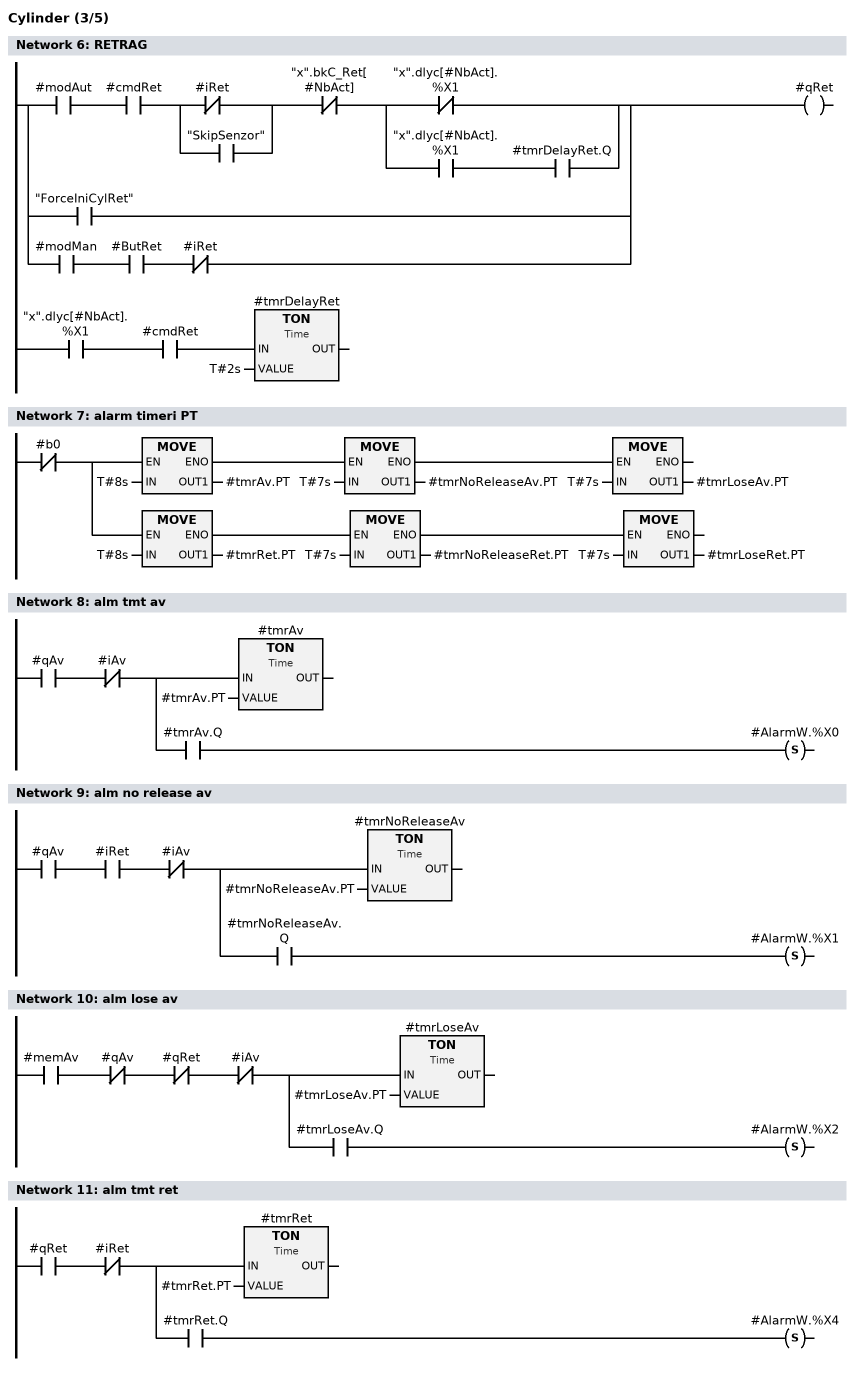
   #qRet := (#modAut AND #cmdRet AND (NOT #iRet OR "SkipSenzor") AND NOT "x".bkC_Ret[#NbAct] AND (NOT "x".dlyc[#NbAct].%X1 OR ("x".dlyc[#NbAct].%X1 AND #tmrDelayRet.Q))) OR "ForceIniCylRet" OR (#modMan AND #ButRet AND NOT #iRet);
   #tmrDelayRet.TON(IN := "x".dlyc[#NbAct].%X1 AND #cmdRet, PT := T#2s);   // TON coil
END_REGION

REGION Network 7: alarm timeri PT
   RUNG wire#powerrail
      I_Contact( #b0 )
      wire#w1
      Move(in := T#8s, out1 => #tmrAv.PT)
      Move(in := T#7s, out1 => #tmrNoReleaseAv.PT)
      Move(in := T#7s, out1 => #tmrLoseAv.PT)
   END_RUNG
   RUNG wire#w1
      Move(in := T#8s, out1 => #tmrRet.PT)
      Move(in := T#7s, out1 => #tmrNoReleaseRet.PT)
      Move(in := T#7s, out1 => #tmrLoseRet.PT)
   END_RUNG
   // the same network as SCL:
   IF NOT #b0 THEN
       #tmrAv.PT := T#8s;
       #tmrNoReleaseAv.PT := T#7s;
       #tmrLoseAv.PT := T#7s;
       #tmrRet.PT := T#8s;
       #tmrNoReleaseRet.PT := T#7s;
       #tmrLoseRet.PT := T#7s;
   END_IF;
END_REGION

REGION Network 8: alm tmt av
   #_w1 := #qAv AND NOT #iAv;
   #tmrAv.TON(IN := #_w1, PT := #tmrAv.PT);   // TON coil
   IF #_w1 AND #tmrAv.Q THEN #AlarmW.%X0 := TRUE; END_IF;
END_REGION

REGION Network 9: alm no release av
   #_w1 := #qAv AND #iRet AND NOT #iAv;
   #tmrNoReleaseAv.TON(IN := #_w1, PT := #tmrNoReleaseAv.PT);   // TON coil
   IF #_w1 AND #tmrNoReleaseAv.Q THEN #AlarmW.%X1 := TRUE; END_IF;
END_REGION

REGION Network 10: alm lose av
   #_w1 := #memAv AND NOT #qAv AND NOT #qRet AND NOT #iAv;
   #tmrLoseAv.TON(IN := #_w1, PT := #tmrLoseAv.PT);   // TON coil
   IF #_w1 AND #tmrLoseAv.Q THEN #AlarmW.%X2 := TRUE; END_IF;
END_REGION

REGION Network 11: alm tmt ret
   #_w1 := #qRet AND NOT #iRet;
   #tmrRet.TON(IN := #_w1, PT := #tmrRet.PT);   // TON coil
   IF #_w1 AND #tmrRet.Q THEN #AlarmW.%X4 := TRUE; END_IF;
END_REGION

REGION Network 12: alm no release ret
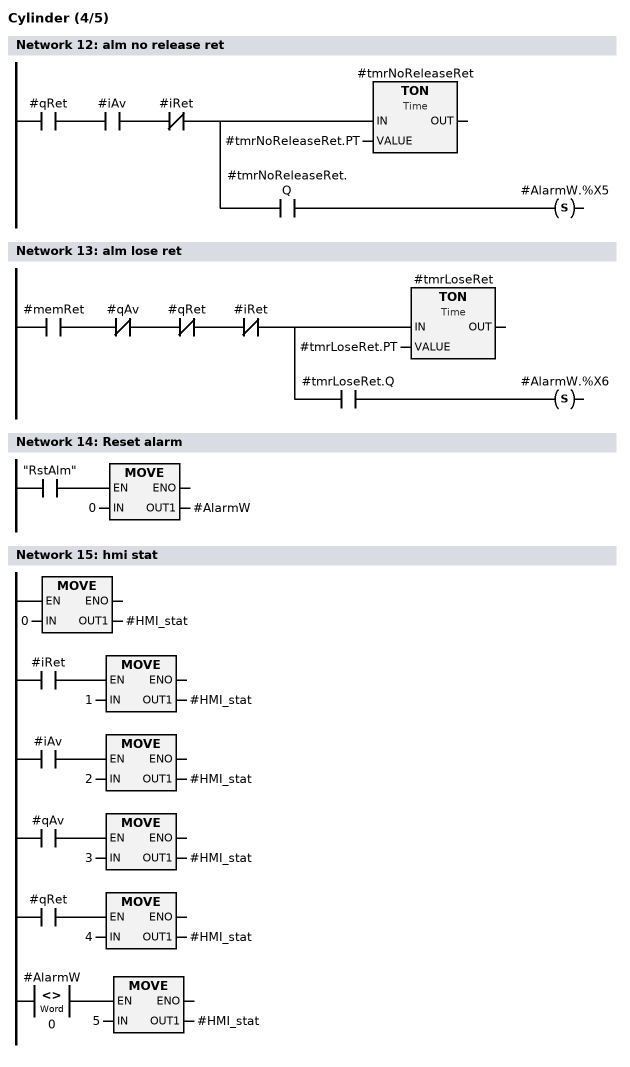
   #_w1 := #qRet AND #iAv AND NOT #iRet;
   #tmrNoReleaseRet.TON(IN := #_w1, PT := #tmrNoReleaseRet.PT);   // TON coil
   IF #_w1 AND #tmrNoReleaseRet.Q THEN #AlarmW.%X5 := TRUE; END_IF;
END_REGION

REGION Network 13: alm lose ret
   #_w1 := #memRet AND NOT #qAv AND NOT #qRet AND NOT #iRet;
   #tmrLoseRet.TON(IN := #_w1, PT := #tmrLoseRet.PT);   // TON coil
   IF #_w1 AND #tmrLoseRet.Q THEN #AlarmW.%X6 := TRUE; END_IF;
END_REGION

REGION Network 14: Reset alarm
   RUNG wire#powerrail
      Contact( "RstAlm" )
      Move(in := 0, out1 => #AlarmW)
   END_RUNG
   // the same network as SCL:
   IF "RstAlm" THEN #AlarmW := 0; END_IF;
END_REGION

REGION Network 15: hmi stat
   RUNG wire#powerrail
      Move(in := 0, out1 => #HMI_stat)
   END_RUNG
   RUNG wire#powerrail
      Contact( #iRet )
      Move(in := 1, out1 => #HMI_stat)
   END_RUNG
   RUNG wire#powerrail
      Contact( #iAv )
      Move(in := 2, out1 => #HMI_stat)
   END_RUNG
   RUNG wire#powerrail
      Contact( #qAv )
      Move(in := 3, out1 => #HMI_stat)
   END_RUNG
   RUNG wire#powerrail
      Contact( #qRet )
      Move(in := 4, out1 => #HMI_stat)
   END_RUNG
   RUNG wire#powerrail
      { S7_Templates := "SrcType := Word" } NE_Contact(in1 := #AlarmW, in2 := 0)
      Move(in := 5, out1 => #HMI_stat)
   END_RUNG
   // the same network as SCL:
   #HMI_stat := 0;
   IF #iRet THEN #HMI_stat := 1; END_IF;
   IF #iAv THEN #HMI_stat := 2; END_IF;
   IF #qAv THEN #HMI_stat := 3; END_IF;
   IF #qRet THEN #HMI_stat := 4; END_IF;
   IF #AlarmW <> 0 THEN #HMI_stat := 5; END_IF;
END_REGION

REGION Network 16: hmi man
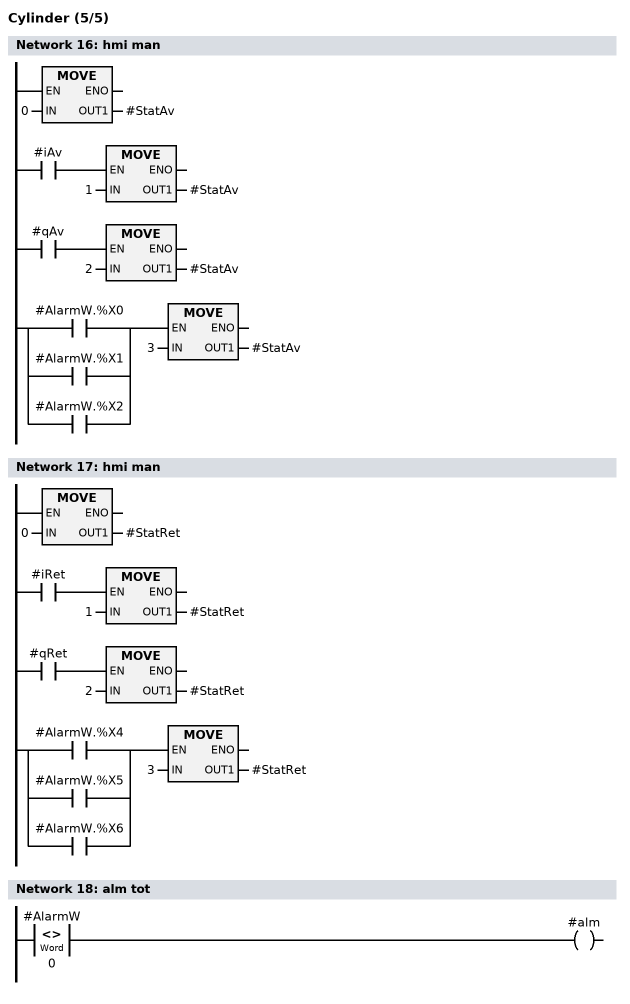
   RUNG wire#powerrail
      Move(in := 0, out1 => #StatAv)
   END_RUNG
   RUNG wire#powerrail
      Contact( #iAv )
      Move(in := 1, out1 => #StatAv)
   END_RUNG
   RUNG wire#powerrail
      Contact( #qAv )
      Move(in := 2, out1 => #StatAv)
   END_RUNG
   RUNG wire#powerrail
      Contact( #AlarmW.%X0 )
      wire#w1
      Move(in := 3, out1 => #StatAv)
   END_RUNG
   RUNG wire#powerrail
      Contact( #AlarmW.%X1 )
   END_RUNG wire#w1
   RUNG wire#powerrail
      Contact( #AlarmW.%X2 )
   END_RUNG wire#w1
   // the same network as SCL:
   #StatAv := 0;
   IF #iAv THEN #StatAv := 1; END_IF;
   IF #qAv THEN #StatAv := 2; END_IF;
   IF #AlarmW.%X0 OR #AlarmW.%X1 OR #AlarmW.%X2 THEN #StatAv := 3; END_IF;
END_REGION

REGION Network 17: hmi man
   RUNG wire#powerrail
      Move(in := 0, out1 => #StatRet)
   END_RUNG
   RUNG wire#powerrail
      Contact( #iRet )
      Move(in := 1, out1 => #StatRet)
   END_RUNG
   RUNG wire#powerrail
      Contact( #qRet )
      Move(in := 2, out1 => #StatRet)
   END_RUNG
   RUNG wire#powerrail
      Contact( #AlarmW.%X4 )
      wire#w1
      Move(in := 3, out1 => #StatRet)
   END_RUNG
   RUNG wire#powerrail
      Contact( #AlarmW.%X5 )
   END_RUNG wire#w1
   RUNG wire#powerrail
      Contact( #AlarmW.%X6 )
   END_RUNG wire#w1
   // the same network as SCL:
   #StatRet := 0;
   IF #iRet THEN #StatRet := 1; END_IF;
   IF #qRet THEN #StatRet := 2; END_IF;
   IF #AlarmW.%X4 OR #AlarmW.%X5 OR #AlarmW.%X6 THEN #StatRet := 3; END_IF;
END_REGION

REGION Network 18: alm tot
   RUNG wire#powerrail
      { S7_Templates := "SrcType := Word" } NE_Contact(in1 := #AlarmW, in2 := 0)
      Coil( #alm )
   END_RUNG
   // the same network as SCL:
   #alm := #AlarmW <> 0;
END_REGION
END_FUNCTION_BLOCK

FUNCTION_BLOCK "FB_Outputs"   // FB8, LAD
{ S7_Optimized_Access := 'TRUE' }
VERSION : 0.1
   VAR
      Centror_A : "Cylinder";
      Centror_B : "Cylinder";
      CilindruVerticalStacker : "Cylinder";
      FurcaStacker : "Cylinder";
      CilindruVerticalStacker_New : "Cylinder";
      FurcaStacker_New : "Cylinder";
      stoper1 : "Cylinder";
      stoper2 : "Cylinder";
      St_Urc_Jos_Sus : Bool;
      St_Urc_Jos_Mijloc : Bool;
      St_Urc_Mijloc_Sus : Bool;
      St_Cobor_Sus_Jos : Bool;
      St_Cobor_Sus_Mijloc : Bool;
      St_Cobor_Mijloc_jos : Bool;
      DSt_Urc_Jos_Sus : Bool;
      DSt_Urc_Jos_Mijloc : Bool;
      DSt_Urc_Mijloc_Sus : Bool;
      DSt_Cobor_Sus_Jos : Bool;
      DSt_Cobor_Sus_Mijloc : Bool;
      DSt_Cobor_Mijloc_jos : Bool;
      StopReqUp1 : Bool;
      StopReqDn1 : Bool;
      StopReqUp2 : Bool;
      StopReqDn2 : Bool;
      S_Alm_Stack_Up : Word;
      S_Alm_Stack_Mid : Word;
      S_Alm_Stack_Dwn : Word;
      SN_Alm_Stack_Up : Word;
      SN_Alm_Stack_Mid : Word;
      SN_Alm_Stack_Dwn : Word;
      Alm_tim : Array[1..9] of IEC_TIMER;
   END_VAR
   VAR_TEMP
      "tmp_Comanda furca extinsa" : Bool;
      "tmp_Comanda furca retrasa" : Bool;
      StopCmd1 : Bool;
      StopCmd2 : Bool;
   END_VAR
BEGIN

REGION Network 1: Stacker : Pasi ridicare coborare
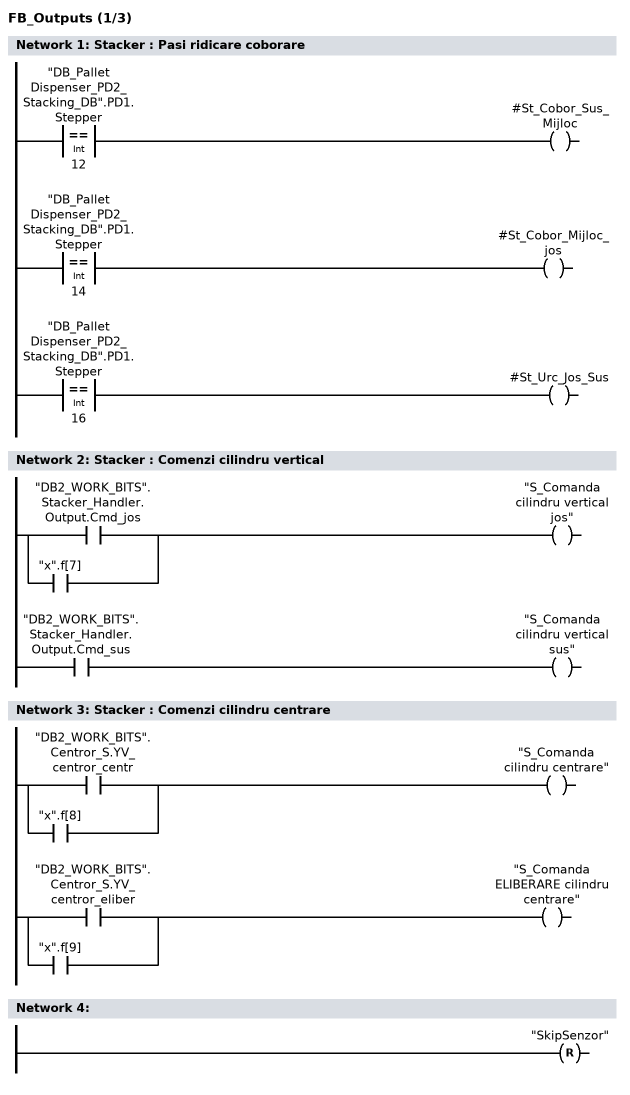
   RUNG wire#powerrail
      { S7_Templates := "SrcType := Int" } EQ_Contact(in1 := "DB_PalletDispenser_PD2_Stacking_DB".PD1.Stepper, in2 := 12)
      Coil( #St_Cobor_Sus_Mijloc )
   END_RUNG
   RUNG wire#powerrail
      { S7_Templates := "SrcType := Int" } EQ_Contact(in1 := "DB_PalletDispenser_PD2_Stacking_DB".PD1.Stepper, in2 := 14)
      Coil( #St_Cobor_Mijloc_jos )
   END_RUNG
   RUNG wire#powerrail
      { S7_Templates := "SrcType := Int" } EQ_Contact(in1 := "DB_PalletDispenser_PD2_Stacking_DB".PD1.Stepper, in2 := 16)
      Coil( #St_Urc_Jos_Sus )
   END_RUNG
   // the same network as SCL:
   #St_Cobor_Sus_Mijloc := "DB_PalletDispenser_PD2_Stacking_DB".PD1.Stepper = 12;
   #St_Cobor_Mijloc_jos := "DB_PalletDispenser_PD2_Stacking_DB".PD1.Stepper = 14;
   #St_Urc_Jos_Sus := "DB_PalletDispenser_PD2_Stacking_DB".PD1.Stepper = 16;
END_REGION

REGION Network 2: Stacker : Comenzi cilindru vertical
   RUNG wire#powerrail
      Contact( "DB2_WORK_BITS".Stacker_Handler.Output.Cmd_jos )
      wire#w1
      Coil( "S_Comanda cilindru vertical jos" )
   END_RUNG
   RUNG wire#powerrail
      Contact( "x".f[7] )
   END_RUNG wire#w1
   RUNG wire#powerrail
      Contact( "DB2_WORK_BITS".Stacker_Handler.Output.Cmd_sus )
      Coil( "S_Comanda cilindru vertical sus" )
   END_RUNG
   // the same network as SCL:
   "S_Comanda cilindru vertical jos" := "DB2_WORK_BITS".Stacker_Handler.Output.Cmd_jos OR "x".f[7];
   "S_Comanda cilindru vertical sus" := "DB2_WORK_BITS".Stacker_Handler.Output.Cmd_sus;
END_REGION

REGION Network 3: Stacker : Comenzi cilindru centrare
   RUNG wire#powerrail
      Contact( "DB2_WORK_BITS".Centror_S.YV_centror_centr )
      wire#w1
      Coil( "S_Comanda cilindru centrare" )
   END_RUNG
   RUNG wire#powerrail
      Contact( "x".f[8] )
   END_RUNG wire#w1
   RUNG wire#powerrail
      Contact( "DB2_WORK_BITS".Centror_S.YV_centror_eliber )
      wire#w2
      Coil( "S_Comanda ELIBERARE cilindru centrare" )
   END_RUNG
   RUNG wire#powerrail
      Contact( "x".f[9] )
   END_RUNG wire#w2
   // the same network as SCL:
   "S_Comanda cilindru centrare" := "DB2_WORK_BITS".Centror_S.YV_centror_centr OR "x".f[8];
   "S_Comanda ELIBERARE cilindru centrare" := "DB2_WORK_BITS".Centror_S.YV_centror_eliber OR "x".f[9];
END_REGION

REGION Network 4
   RUNG wire#powerrail
      R_Coil( "SkipSenzor" )
   END_RUNG
   // the same network as SCL:
   "SkipSenzor" := FALSE;
END_REGION

REGION Network 5: Stacker : Apelare cilindru furca stacker
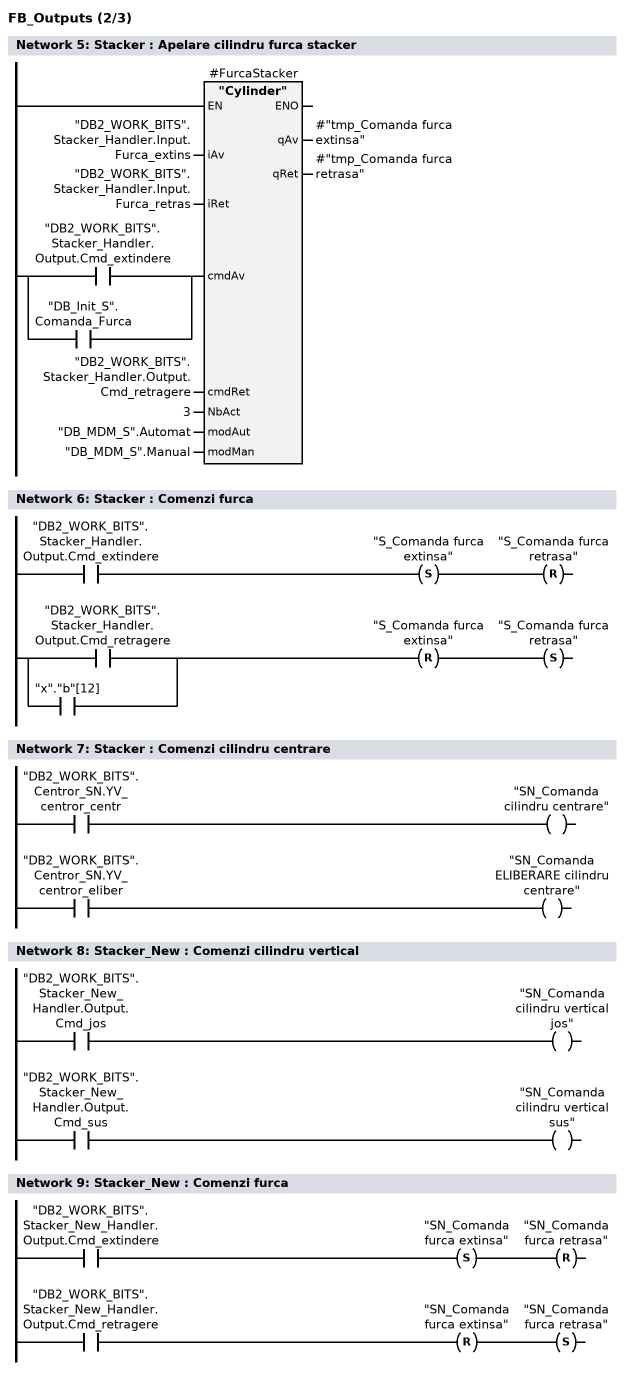
   RUNG wire#powerrail
      #FurcaStacker(cmdAv := wire#w1, iAv := "DB2_WORK_BITS".Stacker_Handler.Input.Furca_extins, iRet := "DB2_WORK_BITS".Stacker_Handler.Input.Furca_retras, cmdRet := "DB2_WORK_BITS".Stacker_Handler.Output.Cmd_retragere, NbAct := 3, modAut := "DB_MDM_S".Automat, modMan := "DB_MDM_S".Manual, qAv => #"tmp_Comanda furca extinsa", qRet => #"tmp_Comanda furca retrasa")
   END_RUNG
   RUNG wire#powerrail
      Contact( "DB2_WORK_BITS".Stacker_Handler.Output.Cmd_extindere )
   END_RUNG wire#w1
   RUNG wire#powerrail
      Contact( "DB_Init_S".Comanda_Furca )
   END_RUNG wire#w1
   // the same network as SCL:
   #FurcaStacker(iAv := "DB2_WORK_BITS".Stacker_Handler.Input.Furca_extins,   // "Cylinder"
                 iRet := "DB2_WORK_BITS".Stacker_Handler.Input.Furca_retras,
                 cmdAv := "DB2_WORK_BITS".Stacker_Handler.Output.Cmd_extindere OR "DB_Init_S".Comanda_Furca,
                 cmdRet := "DB2_WORK_BITS".Stacker_Handler.Output.Cmd_retragere,
                 NbAct := 3,
                 modAut := "DB_MDM_S".Automat,
                 modMan := "DB_MDM_S".Manual,
                 qAv => #"tmp_Comanda furca extinsa",
                 qRet => #"tmp_Comanda furca retrasa");
END_REGION

REGION Network 6: Stacker : Comenzi furca
   RUNG wire#powerrail
      Contact( "DB2_WORK_BITS".Stacker_Handler.Output.Cmd_extindere )
      S_Coil( "S_Comanda furca extinsa" )
      R_Coil( "S_Comanda furca retrasa" )
   END_RUNG
   RUNG wire#powerrail
      Contact( "DB2_WORK_BITS".Stacker_Handler.Output.Cmd_retragere )
      wire#w1
      R_Coil( "S_Comanda furca extinsa" )
      S_Coil( "S_Comanda furca retrasa" )
   END_RUNG
   RUNG wire#powerrail
      Contact( "x"."b"[12] )
   END_RUNG wire#w1
   // the same network as SCL:
   IF "DB2_WORK_BITS".Stacker_Handler.Output.Cmd_extindere THEN
       "S_Comanda furca extinsa" := TRUE;
       "S_Comanda furca retrasa" := FALSE;
   END_IF;
   IF "DB2_WORK_BITS".Stacker_Handler.Output.Cmd_retragere OR "x"."b"[12] THEN
       "S_Comanda furca extinsa" := FALSE;
       "S_Comanda furca retrasa" := TRUE;
   END_IF;
END_REGION

REGION Network 7: Stacker : Comenzi cilindru centrare
   RUNG wire#powerrail
      Contact( "DB2_WORK_BITS".Centror_SN.YV_centror_centr )
      Coil( "SN_Comanda cilindru centrare" )
   END_RUNG
   RUNG wire#powerrail
      Contact( "DB2_WORK_BITS".Centror_SN.YV_centror_eliber )
      Coil( "SN_Comanda ELIBERARE cilindru centrare" )
   END_RUNG
   // the same network as SCL:
   "SN_Comanda cilindru centrare" := "DB2_WORK_BITS".Centror_SN.YV_centror_centr;
   "SN_Comanda ELIBERARE cilindru centrare" := "DB2_WORK_BITS".Centror_SN.YV_centror_eliber;
END_REGION

REGION Network 8: Stacker_New : Comenzi cilindru vertical
   RUNG wire#powerrail
      Contact( "DB2_WORK_BITS".Stacker_New_Handler.Output.Cmd_jos )
      Coil( "SN_Comanda cilindru vertical jos" )
   END_RUNG
   RUNG wire#powerrail
      Contact( "DB2_WORK_BITS".Stacker_New_Handler.Output.Cmd_sus )
      Coil( "SN_Comanda cilindru vertical sus" )
   END_RUNG
   // the same network as SCL:
   "SN_Comanda cilindru vertical jos" := "DB2_WORK_BITS".Stacker_New_Handler.Output.Cmd_jos;
   "SN_Comanda cilindru vertical sus" := "DB2_WORK_BITS".Stacker_New_Handler.Output.Cmd_sus;
END_REGION

REGION Network 9: Stacker_New : Comenzi furca
   RUNG wire#powerrail
      Contact( "DB2_WORK_BITS".Stacker_New_Handler.Output.Cmd_extindere )
      S_Coil( "SN_Comanda furca extinsa" )
      R_Coil( "SN_Comanda furca retrasa" )
   END_RUNG
   RUNG wire#powerrail
      Contact( "DB2_WORK_BITS".Stacker_New_Handler.Output.Cmd_retragere )
      R_Coil( "SN_Comanda furca extinsa" )
      S_Coil( "SN_Comanda furca retrasa" )
   END_RUNG
   // the same network as SCL:
   IF "DB2_WORK_BITS".Stacker_New_Handler.Output.Cmd_extindere THEN
       "SN_Comanda furca extinsa" := TRUE;
       "SN_Comanda furca retrasa" := FALSE;
   END_IF;
   IF "DB2_WORK_BITS".Stacker_New_Handler.Output.Cmd_retragere THEN
       "SN_Comanda furca extinsa" := FALSE;
       "SN_Comanda furca retrasa" := TRUE;
   END_IF;
END_REGION

REGION Network 10: Stacker_New : Apelare cilindru furca
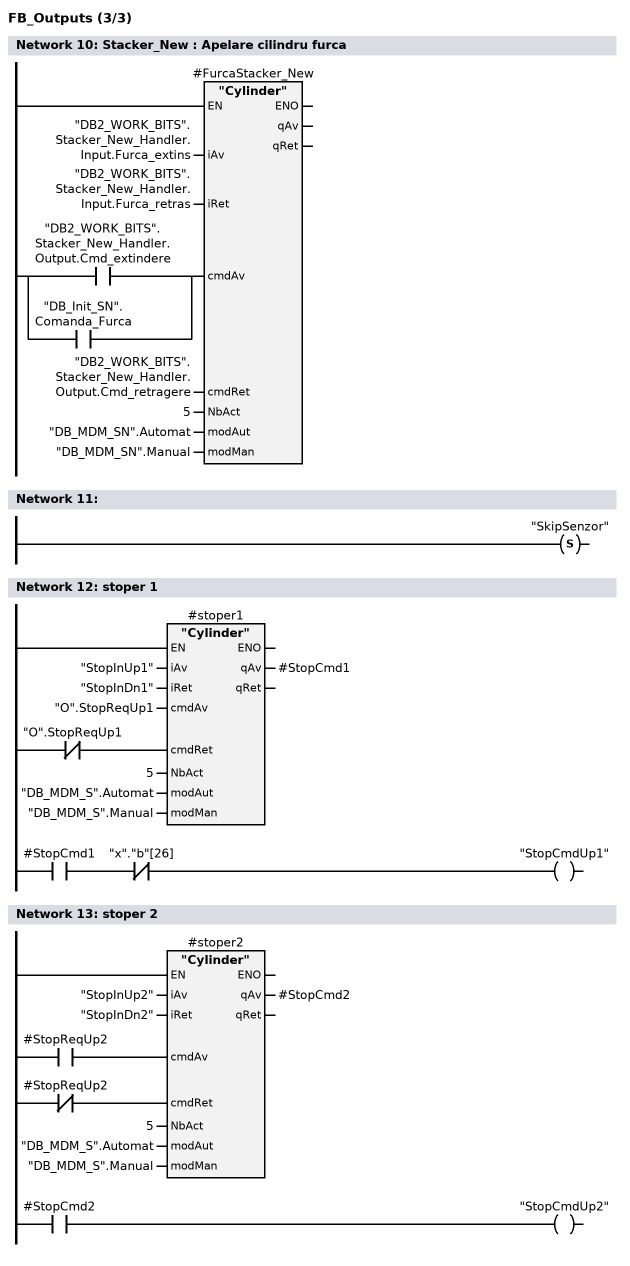
   RUNG wire#powerrail
      #FurcaStacker_New(cmdAv := wire#w1, iAv := "DB2_WORK_BITS".Stacker_New_Handler.Input.Furca_extins, iRet := "DB2_WORK_BITS".Stacker_New_Handler.Input.Furca_retras, cmdRet := "DB2_WORK_BITS".Stacker_New_Handler.Output.Cmd_retragere, NbAct := 5, modAut := "DB_MDM_SN".Automat, modMan := "DB_MDM_SN".Manual, qAv =>, qRet =>)
   END_RUNG
   RUNG wire#powerrail
      Contact( "DB2_WORK_BITS".Stacker_New_Handler.Output.Cmd_extindere )
   END_RUNG wire#w1
   RUNG wire#powerrail
      Contact( "DB_Init_SN".Comanda_Furca )
   END_RUNG wire#w1
   // the same network as SCL:
   #FurcaStacker_New(iAv := "DB2_WORK_BITS".Stacker_New_Handler.Input.Furca_extins,   // "Cylinder"
                     iRet := "DB2_WORK_BITS".Stacker_New_Handler.Input.Furca_retras,
                     cmdAv := "DB2_WORK_BITS".Stacker_New_Handler.Output.Cmd_extindere OR "DB_Init_SN".Comanda_Furca,
                     cmdRet := "DB2_WORK_BITS".Stacker_New_Handler.Output.Cmd_retragere,
                     NbAct := 5,
                     modAut := "DB_MDM_SN".Automat,
                     modMan := "DB_MDM_SN".Manual);
END_REGION

REGION Network 11
   RUNG wire#powerrail
      S_Coil( "SkipSenzor" )
   END_RUNG
   // the same network as SCL:
   "SkipSenzor" := TRUE;
END_REGION

REGION Network 12: stoper 1
   RUNG wire#powerrail
      #stoper1(cmdRet := wire#w1, iAv := "StopInUp1", iRet := "StopInDn1", cmdAv := "O".StopReqUp1, NbAct := 5, modAut := "DB_MDM_S".Automat, modMan := "DB_MDM_S".Manual, qAv => #StopCmd1, qRet =>)
   END_RUNG
   RUNG wire#powerrail
      I_Contact( "O".StopReqUp1 )
   END_RUNG wire#w1
   RUNG wire#powerrail
      Contact( #StopCmd1 )
      I_Contact( "x"."b"[26] )
      Coil( "StopCmdUp1" )
   END_RUNG
   // the same network as SCL:
   #stoper1(iAv := "StopInUp1",   // "Cylinder"
            iRet := "StopInDn1",
            cmdAv := "O".StopReqUp1,
            cmdRet := NOT "O".StopReqUp1,
            NbAct := 5,
            modAut := "DB_MDM_S".Automat,
            modMan := "DB_MDM_S".Manual,
            qAv => #StopCmd1);
   "StopCmdUp1" := #StopCmd1 AND NOT "x"."b"[26];
END_REGION

REGION Network 13: stoper 2
   RUNG wire#powerrail
      #stoper2(cmdAv := wire#w1, cmdRet := wire#w2, iAv := "StopInUp2", iRet := "StopInDn2", NbAct := 5, modAut := "DB_MDM_S".Automat, modMan := "DB_MDM_S".Manual, qAv => #StopCmd2, qRet =>)
   END_RUNG
   RUNG wire#powerrail
      Contact( #StopReqUp2 )
   END_RUNG wire#w1
   RUNG wire#powerrail
      I_Contact( #StopReqUp2 )
   END_RUNG wire#w2
   RUNG wire#powerrail
      Contact( #StopCmd2 )
      Coil( "StopCmdUp2" )
   END_RUNG
   // the same network as SCL:
   #stoper2(iAv := "StopInUp2",   // "Cylinder"
            iRet := "StopInDn2",
            cmdAv := #StopReqUp2,
            cmdRet := NOT #StopReqUp2,
            NbAct := 5,
            modAut := "DB_MDM_S".Automat,
            modMan := "DB_MDM_S".Manual,
            qAv => #StopCmd2);
   "StopCmdUp2" := #StopCmd2;
END_REGION
END_FUNCTION_BLOCK

FUNCTION_BLOCK "FB_MDM"   // FB10, LAD
{ S7_Optimized_Access := 'TRUE' }
VERSION : 0.1
// td -inlocuit biti GEN cu intrari
// td inlocuit biti M.15.4 "Cycle_Run_S" cu bitii  DB.Cycle_Run peste tot in program
   VAR_INPUT
      ButAuto : Bool;
      cndSafe : Bool;
      cndEnergie : Bool;
      Home : Bool;
      ButStartCycle : Bool;
      AlarmStop : Bool;
      ButInit : Bool;
      ButStep : Bool;
      ButStopCycle : Bool;
      G7_Stack : Int;
   END_VAR
   VAR_IN_OUT
      Init_OK : Bool;
      Init_Req : Bool;
   END_VAR
   VAR
      No_Safe : Bool;
      Energie : Bool;
      Manual : Bool;
      Automat : Bool;
      Wait_Start_Cycle : Bool;
      Cycle_Run : Bool;
      Init : Bool;
      Init_Done : Bool;
      Safe : Bool;
      "step" : USInt;
      stepimg : USInt;
      Stepper : Bool;
   END_VAR
   VAR_TEMP   // added for the SCL form of the ladder/FBD networks
      _w1 : Bool;
   END_VAR
BEGIN

REGION Network 1: First cycle
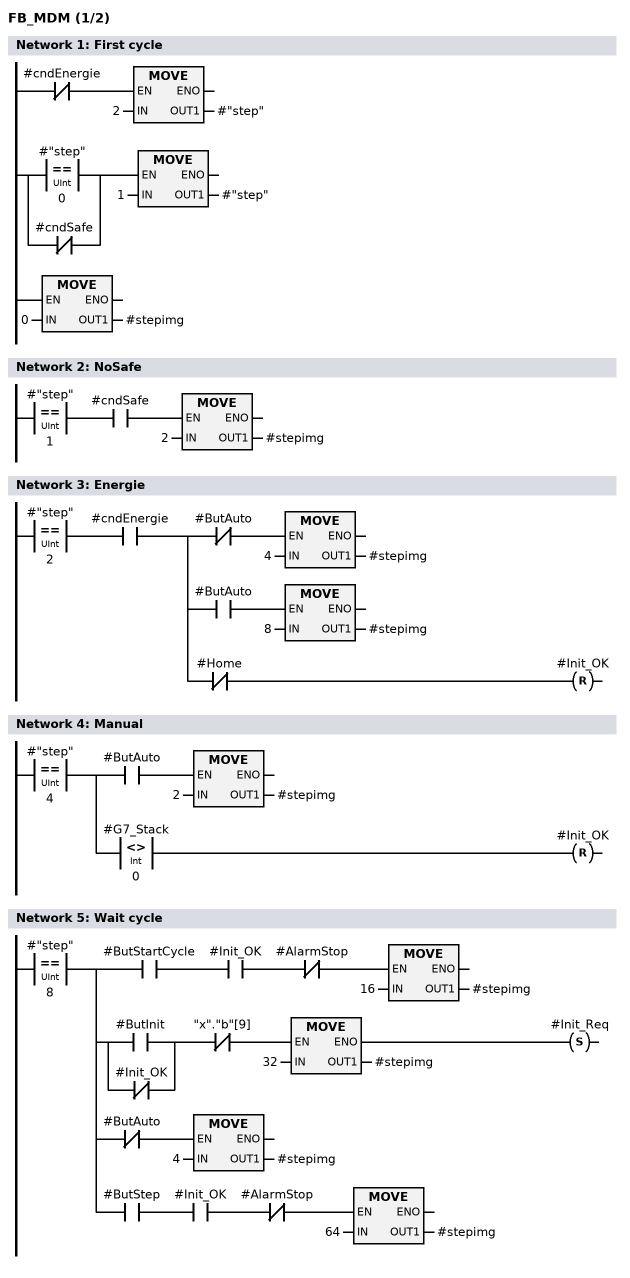
   RUNG wire#powerrail
      I_Contact( #cndEnergie )
      Move(in := 2, out1 => #"step")
   END_RUNG
   RUNG wire#powerrail
      { S7_Templates := "SrcType := UInt" } EQ_Contact(in1 := #"step", in2 := 0)
      wire#w1
      Move(in := 1, out1 => #"step")
   END_RUNG
   RUNG wire#powerrail
      I_Contact( #cndSafe )
   END_RUNG wire#w1
   RUNG wire#powerrail
      Move(in := 0, out1 => #stepimg)
   END_RUNG
   // the same network as SCL:
   IF NOT #cndEnergie THEN #"step" := 2; END_IF;
   IF (#"step" = 0) OR NOT #cndSafe THEN #"step" := 1; END_IF;
   #stepimg := 0;
END_REGION

REGION Network 2: NoSafe
   RUNG wire#powerrail
      { S7_Templates := "SrcType := UInt" } EQ_Contact(in1 := #"step", in2 := 1)
      Contact( #cndSafe )
      Move(in := 2, out1 => #stepimg)
   END_RUNG
   // the same network as SCL:
   IF (#"step" = 1) AND #cndSafe THEN #stepimg := 2; END_IF;
END_REGION

REGION Network 3: Energie
   RUNG wire#powerrail
      { S7_Templates := "SrcType := UInt" } EQ_Contact(in1 := #"step", in2 := 2)
      Contact( #cndEnergie )
      wire#w1
      I_Contact( #ButAuto )
      Move(in := 4, out1 => #stepimg)
   END_RUNG
   RUNG wire#w1
      Contact( #ButAuto )
      Move(in := 8, out1 => #stepimg)
   END_RUNG
   RUNG wire#w1
      I_Contact( #Home )
      R_Coil( #Init_OK )
   END_RUNG
   // the same network as SCL:
   #_w1 := (#"step" = 2) AND #cndEnergie;
   IF #_w1 AND NOT #ButAuto THEN #stepimg := 4; END_IF;
   IF #_w1 AND #ButAuto THEN #stepimg := 8; END_IF;
   IF #_w1 AND NOT #Home THEN #Init_OK := FALSE; END_IF;
END_REGION

REGION Network 4: Manual
   RUNG wire#powerrail
      { S7_Templates := "SrcType := UInt" } EQ_Contact(in1 := #"step", in2 := 4)
      wire#w1
      Contact( #ButAuto )
      Move(in := 2, out1 => #stepimg)
   END_RUNG
   RUNG wire#w1
      { S7_Templates := "SrcType := Int" } NE_Contact(in1 := #G7_Stack, in2 := 0)
      R_Coil( #Init_OK )
   END_RUNG
   // the same network as SCL:
   #_w1 := #"step" = 4;
   IF #_w1 AND #ButAuto THEN #stepimg := 2; END_IF;
   IF #_w1 AND (#G7_Stack <> 0) THEN #Init_OK := FALSE; END_IF;
END_REGION

REGION Network 5: Wait cycle
   RUNG wire#powerrail
      { S7_Templates := "SrcType := UInt" } EQ_Contact(in1 := #"step", in2 := 8)
      wire#w1
      Contact( #ButStartCycle )
      Contact( #Init_OK )
      I_Contact( #AlarmStop )
      Move(in := 16, out1 => #stepimg)
   END_RUNG
   RUNG wire#w1
      Contact( #ButInit )
      wire#w2
      I_Contact( "x"."b"[9] )
      Move(in := 32, out1 => #stepimg)
      S_Coil( #Init_Req )
   END_RUNG
   RUNG wire#w1
      I_Contact( #Init_OK )
   END_RUNG wire#w2
   RUNG wire#w1
      I_Contact( #ButAuto )
      Move(in := 4, out1 => #stepimg)
   END_RUNG
   RUNG wire#w1
      Contact( #ButStep )
      Contact( #Init_OK )
      I_Contact( #AlarmStop )
      Move(in := 64, out1 => #stepimg)
   END_RUNG
   // the same network as SCL:
   #_w1 := #"step" = 8;
   IF #_w1 AND #ButStartCycle AND #Init_OK AND NOT #AlarmStop THEN #stepimg := 16; END_IF;
   IF #_w1 AND (#ButInit OR NOT #Init_OK) AND NOT "x"."b"[9] THEN
       #stepimg := 32;
       #Init_Req := TRUE;
   END_IF;
   IF #_w1 AND NOT #ButAuto THEN #stepimg := 4; END_IF;
   IF #_w1 AND #ButStep AND #Init_OK AND NOT #AlarmStop THEN #stepimg := 64; END_IF;
END_REGION

REGION Network 6: Init
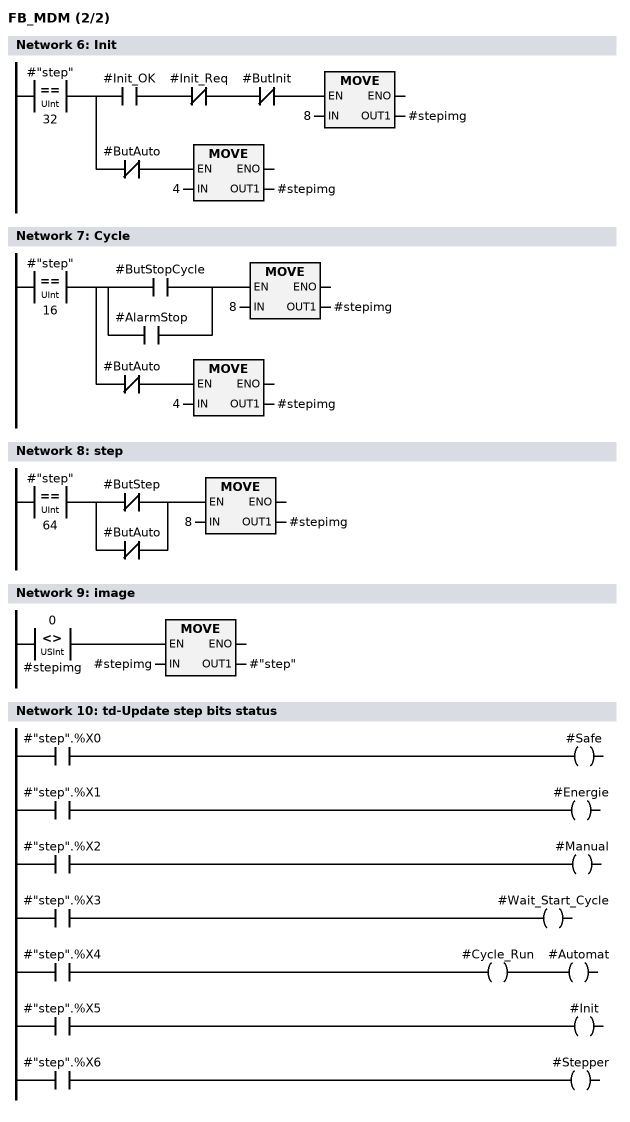
   RUNG wire#powerrail
      { S7_Templates := "SrcType := UInt" } EQ_Contact(in1 := #"step", in2 := 32)
      wire#w1
      Contact( #Init_OK )
      I_Contact( #Init_Req )
      I_Contact( #ButInit )
      Move(in := 8, out1 => #stepimg)
   END_RUNG
   RUNG wire#w1
      I_Contact( #ButAuto )
      Move(in := 4, out1 => #stepimg)
   END_RUNG
   // the same network as SCL:
   #_w1 := #"step" = 32;
   IF #_w1 AND #Init_OK AND NOT #Init_Req AND NOT #ButInit THEN #stepimg := 8; END_IF;
   IF #_w1 AND NOT #ButAuto THEN #stepimg := 4; END_IF;
END_REGION

REGION Network 7: Cycle
   RUNG wire#powerrail
      { S7_Templates := "SrcType := UInt" } EQ_Contact(in1 := #"step", in2 := 16)
      wire#w1
      Contact( #ButStopCycle )
      wire#w2
      Move(in := 8, out1 => #stepimg)
   END_RUNG
   RUNG wire#w1
      Contact( #AlarmStop )
   END_RUNG wire#w2
   RUNG wire#w1
      I_Contact( #ButAuto )
      Move(in := 4, out1 => #stepimg)
   END_RUNG
   // the same network as SCL:
   #_w1 := #"step" = 16;
   IF #_w1 AND (#ButStopCycle OR #AlarmStop) THEN #stepimg := 8; END_IF;
   IF #_w1 AND NOT #ButAuto THEN #stepimg := 4; END_IF;
END_REGION

REGION Network 8: step
   RUNG wire#powerrail
      { S7_Templates := "SrcType := UInt" } EQ_Contact(in1 := #"step", in2 := 64)
      wire#w1
      I_Contact( #ButStep )
      wire#w2
      Move(in := 8, out1 => #stepimg)
   END_RUNG
   RUNG wire#w1
      I_Contact( #ButAuto )
   END_RUNG wire#w2
   // the same network as SCL:
   IF (#"step" = 64) AND (NOT #ButStep OR NOT #ButAuto) THEN #stepimg := 8; END_IF;
END_REGION

REGION Network 9: image
   RUNG wire#powerrail
      { S7_Templates := "SrcType := USInt" } NE_Contact(in1 := 0, in2 := #stepimg)
      Move(in := #stepimg, out1 => #"step")
   END_RUNG
   // the same network as SCL:
   IF 0 <> #stepimg THEN #"step" := #stepimg; END_IF;
END_REGION

REGION Network 10: td-Update step bits status
   RUNG wire#powerrail
      Contact( #"step".%X0 )
      Coil( #Safe )
   END_RUNG
   RUNG wire#powerrail
      Contact( #"step".%X1 )
      Coil( #Energie )
   END_RUNG
   RUNG wire#powerrail
      Contact( #"step".%X2 )
      Coil( #Manual )
   END_RUNG
   RUNG wire#powerrail
      Contact( #"step".%X3 )
      Coil( #Wait_Start_Cycle )
   END_RUNG
   RUNG wire#powerrail
      Contact( #"step".%X4 )
      Coil( #Cycle_Run )
      Coil( #Automat )
   END_RUNG
   RUNG wire#powerrail
      Contact( #"step".%X5 )
      Coil( #Init )
   END_RUNG
   RUNG wire#powerrail
      Contact( #"step".%X6 )
      Coil( #Stepper )
   END_RUNG
   // the same network as SCL:
   #Safe := #"step".%X0;
   #Energie := #"step".%X1;
   #Manual := #"step".%X2;
   #Wait_Start_Cycle := #"step".%X3;
   #Cycle_Run := #"step".%X4;
   #Automat := #"step".%X4;
   #Init := #"step".%X5;
   #Stepper := #"step".%X6;
END_REGION
END_FUNCTION_BLOCK

FUNCTION_BLOCK "simCylinder"   // FB11, LAD
{ S7_Optimized_Access := 'TRUE' }
VERSION : 0.1
   VAR_INPUT
      qAv : Bool;
      qRet : Bool;
   END_VAR
   VAR_OUTPUT
      iAv : Bool;
      iRet : Bool;
   END_VAR
BEGIN

REGION Network 1
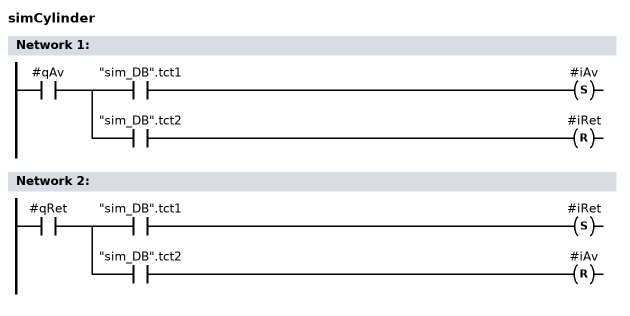
   RUNG wire#powerrail
      Contact( #qAv )
      wire#w1
      Contact( "sim_DB".tct1 )
      S_Coil( #iAv )
   END_RUNG
   RUNG wire#w1
      Contact( "sim_DB".tct2 )
      R_Coil( #iRet )
   END_RUNG
   // the same network as SCL:
   IF #qAv AND "sim_DB".tct1 THEN #iAv := TRUE; END_IF;
   IF #qAv AND "sim_DB".tct2 THEN #iRet := FALSE; END_IF;
END_REGION

REGION Network 2
   RUNG wire#powerrail
      Contact( #qRet )
      wire#w1
      Contact( "sim_DB".tct1 )
      S_Coil( #iRet )
   END_RUNG
   RUNG wire#w1
      Contact( "sim_DB".tct2 )
      R_Coil( #iAv )
   END_RUNG
   // the same network as SCL:
   IF #qRet AND "sim_DB".tct1 THEN #iRet := TRUE; END_IF;
   IF #qRet AND "sim_DB".tct2 THEN #iAv := FALSE; END_IF;
END_REGION
END_FUNCTION_BLOCK

FUNCTION_BLOCK "StaCall"   // FB12, LAD
{ S7_Optimized_Access := 'TRUE' }
VERSION : 0.1
   VAR
      f : Array[0..10] of "sta";
      tranzit : Array[0..10] of Bool;
      Range_LS_1 : Bool;
      Range_LS_2 : Bool;
      Range_LS_3 : Bool;
      PrezPalStackLength : Bool;
      PrezPalStackAnyLength : Bool;
      PrezPalStackAny : Bool;
      DeliveryStack : Bool;
      StivStat : USInt;
      nAc : USInt;
      tmrSnzCentr : TON_TIME;
      tmr : Array[0..8] of IEC_TIMER;
   END_VAR
   VAR_TEMP
      to_ce : Bool;
      to_cm : Bool;
      cmdLiftUpO : Bool;
      tranzit12 : Bool;
   END_VAR
   VAR CONSTANT
      _nop0 : Int := 0;
      _op1 : Int := 1;
      _op2 : Int := 2;
      _cen : Int := 3;
      _stack : Int := 4;
      _evac : Int := 5;
      _nop : Int := 6;
   END_VAR
   VAR_TEMP   // added for the SCL form of the ladder/FBD networks
      _w1 : Bool;
      _w2 : Bool;
      _w3 : Bool;
   END_VAR
BEGIN

REGION Network 1: Force init
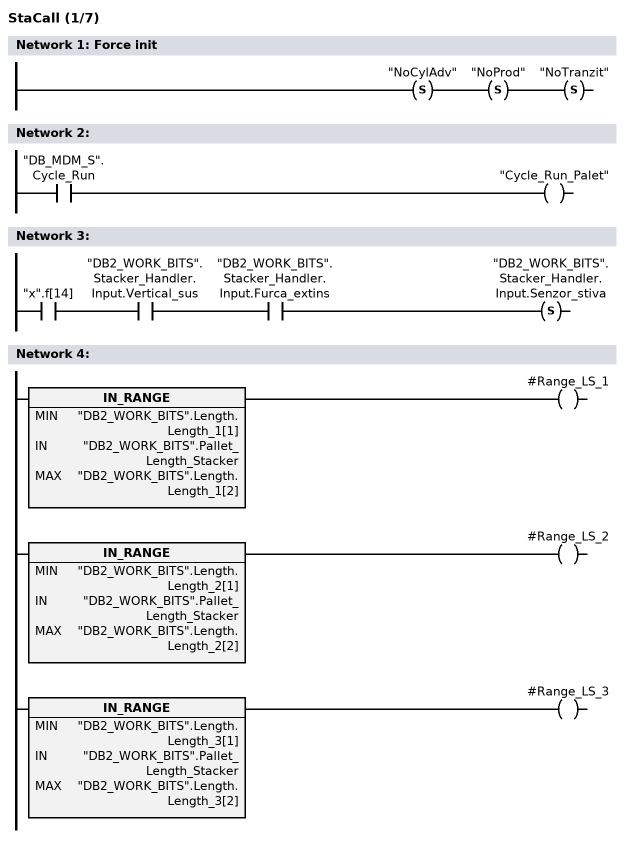
   RUNG wire#powerrail
      S_Coil( "NoCylAdv" )
      S_Coil( "NoProd" )
      S_Coil( "NoTranzit" )
   END_RUNG
   // the same network as SCL:
   "NoCylAdv" := TRUE;
   "NoProd" := TRUE;
   "NoTranzit" := TRUE;
END_REGION

REGION Network 2
   RUNG wire#powerrail
      Contact( "DB_MDM_S".Cycle_Run )
      Coil( "Cycle_Run_Palet" )
   END_RUNG
   // the same network as SCL:
   "Cycle_Run_Palet" := "DB_MDM_S".Cycle_Run;
END_REGION

REGION Network 3
   RUNG wire#powerrail
      Contact( "x".f[14] )
      Contact( "DB2_WORK_BITS".Stacker_Handler.Input.Vertical_sus )
      Contact( "DB2_WORK_BITS".Stacker_Handler.Input.Furca_extins )
      S_Coil( "DB2_WORK_BITS".Stacker_Handler.Input.Senzor_stiva )
   END_RUNG
   // the same network as SCL:
   IF "x".f[14] AND "DB2_WORK_BITS".Stacker_Handler.Input.Vertical_sus AND "DB2_WORK_BITS".Stacker_Handler.Input.Furca_extins THEN
       "DB2_WORK_BITS".Stacker_Handler.Input.Senzor_stiva := TRUE;
   END_IF;
END_REGION

REGION Network 4
   RUNG wire#powerrail
      { S7_Templates := "SrcType := Int" } InRange(min := "DB2_WORK_BITS".Length.Length_1[1], in := "DB2_WORK_BITS".Pallet_Length_Stacker, max := "DB2_WORK_BITS".Length.Length_1[2])
      Coil( #Range_LS_1 )
   END_RUNG
   RUNG wire#powerrail
      { S7_Templates := "SrcType := Int" } InRange(min := "DB2_WORK_BITS".Length.Length_2[1], in := "DB2_WORK_BITS".Pallet_Length_Stacker, max := "DB2_WORK_BITS".Length.Length_2[2])
      Coil( #Range_LS_2 )
   END_RUNG
   RUNG wire#powerrail
      { S7_Templates := "SrcType := Int" } InRange(min := "DB2_WORK_BITS".Length.Length_3[1], in := "DB2_WORK_BITS".Pallet_Length_Stacker, max := "DB2_WORK_BITS".Length.Length_3[2])
      Coil( #Range_LS_3 )
   END_RUNG
   // the same network as SCL:
   #Range_LS_1 := ("DB2_WORK_BITS".Length.Length_1[1] <= "DB2_WORK_BITS".Pallet_Length_Stacker) AND ("DB2_WORK_BITS".Pallet_Length_Stacker <= "DB2_WORK_BITS".Length.Length_1[2]);
   #Range_LS_2 := ("DB2_WORK_BITS".Length.Length_2[1] <= "DB2_WORK_BITS".Pallet_Length_Stacker) AND ("DB2_WORK_BITS".Pallet_Length_Stacker <= "DB2_WORK_BITS".Length.Length_2[2]);
   #Range_LS_3 := ("DB2_WORK_BITS".Length.Length_3[1] <= "DB2_WORK_BITS".Pallet_Length_Stacker) AND ("DB2_WORK_BITS".Pallet_Length_Stacker <= "DB2_WORK_BITS".Length.Length_3[2]);
END_REGION

REGION Network 5: 1 Op1
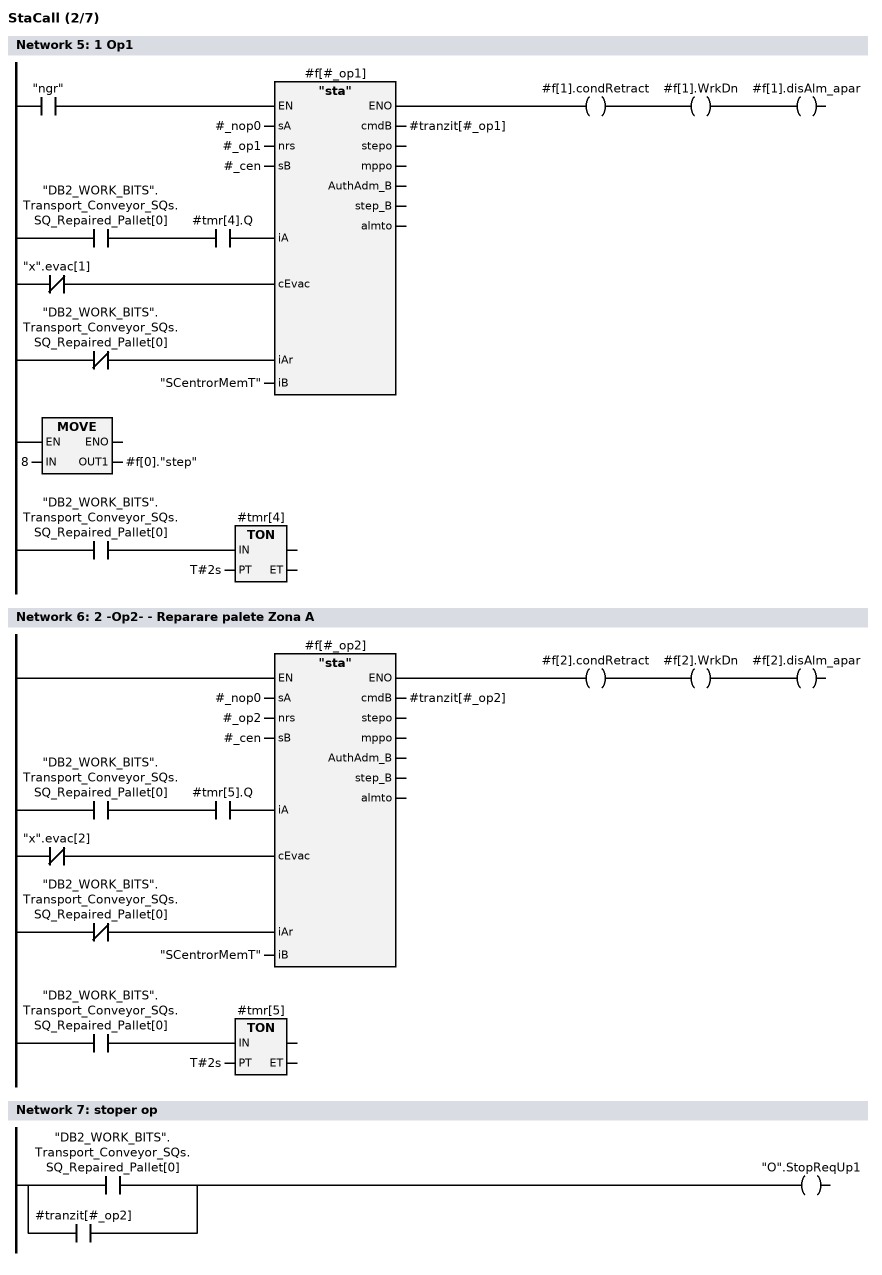
   #f[#_op1](EN := "ngr",   // "sta"
             sA := #_nop0,
             nrs := #_op1,
             sB := #_cen,
             iA := "DB2_WORK_BITS".Transport_Conveyor_SQs.SQ_Repaired_Pallet[0] AND #tmr[4].Q,
             cEvac := NOT "x".evac[1],
             iAr := NOT "DB2_WORK_BITS".Transport_Conveyor_SQs.SQ_Repaired_Pallet[0],
             iB := "SCentrorMemT",
             cmdB => #tranzit[#_op1],
             ENO => #_w1);
   #f[1].condRetract := #_w1;
   #f[1].WrkDn := #_w1;
   #f[1].disAlm_apar := #_w1;
   #f[0]."step" := 8;
   #tmr[4].TON(IN := "DB2_WORK_BITS".Transport_Conveyor_SQs.SQ_Repaired_Pallet[0], PT := T#2s);
END_REGION

